
     // Popup for device diagnostics
     IF ((#hmiData.ioSlotDiagnosticsLoaded = TRUE)
       AND (#statActDeviceOfScreen >= 1)
       AND (#statActDeviceOfScreen <= "USERDIAG_DEVICES_PER_SCREEN_UPPER_LIM"))
     THEN
       #tempDeviceIndex := UINT_TO_INT(#hmiData.actIOSystemData.actIODeviceNumbers[#statActDeviceOfScreen]);
       #hmiData.actDeviceName := #ioSystemData[#statActIOSystem].devices[#tempDeviceIndex].name;
       #hmiData.actDeviceNumber := #ioSystemData[#statActIOSystem].devices[#tempDeviceIndex].number;
       #hmiData.actIPAddress := #ioSystemData[#statActIOSystem].devices[#tempDeviceIndex].ipAddress;

       FOR #tempIndex := 0 TO "USERDIAG_SLOTS_PER_SCREEN_UPPER_LIM" DO
         IF (#tempIndex <= "USERDIAG_SLOTS_PER_DEVICE_UPPER_LIM")
         THEN
           #hmiData.actIOSystemData.actDeviceSlotsUsed[#tempIndex] := (#ioSystemData[#statActIOSystem].devices[#tempDeviceIndex].slots[#tempIndex].configured);
           #hmiData.actIOSystemData.actDeviceSlotsState[#tempIndex] := #ioSystemData[#statActIOSystem].devices[#tempDeviceIndex].slots[#tempIndex].state;
         ELSE
           #hmiData.actIOSystemData.actDeviceSlotsUsed[#tempIndex] := FALSE;
           #hmiData.actIOSystemData.actDeviceSlotsState[#tempIndex] := 0;
         END_IF;
       END_FOR;
     END_IF;
     //===============================================================================================================
     // Colors the button, which switches the actual Screen of Devices in case of faulty Device is on different Screen
     //===============================================================================================================
     #tempIndex := 1;
     #tempErrorStateLower := FALSE;
     // Check if devices before the shown in actual Screen are faulty
     WHILE (#tempIndex <= (#hmiData.actIOSystemData.actIODeviceNumbers[1] - 1))
     DO
       IF ((#ioSystemData[#statActIOSystem].devices[#tempIndex].state = #STATE_FAULT)
         OR (#ioSystemData[#statActIOSystem].devices[#tempIndex].state = #STATE_LOST_CON)
         OR (#ioSystemData[#statActIOSystem].devices[#tempIndex].state = #STATE_PROBLEM))
       THEN
         #tempErrorStateLower := TRUE;
       END_IF;
       #tempIndex := #tempIndex + 1;
     END_WHILE;

     #hmiData.errorAtLowerScreen := #tempErrorStateLower;

     #tempIndex := UINT_TO_INT(#hmiData.actIOSystemData.actIODeviceNumbers["USERDIAG_DEVICES_PER_SCREEN_UPPER_LIM"] + 1);
     #tempErrorStateUpper := FALSE;
     // Check if devices after the shown in actual Screen are faulty
     IF (#tempIndex > 1)
     THEN
       WHILE ((#tempIndex <= #ioSystemData[#statActIOSystem].lastDevice))
       DO
         IF ((#ioSystemData[#statActIOSystem].devices[#tempIndex].state = #STATE_FAULT)
           OR (#ioSystemData[#statActIOSystem].devices[#tempIndex].state = #STATE_LOST_CON)
           OR (#ioSystemData[#statActIOSystem].devices[#tempIndex].state = #STATE_PROBLEM))
         THEN
           #tempErrorStateUpper := TRUE;
         END_IF;
         #tempIndex := #tempIndex + 1;
       END_WHILE;
     END_IF;

     #hmiData.errorAtUpperScreen := #tempErrorStateUpper;
     //=============================================================================
     // Check if PLC diagnostics is selected
     //=============================================================================
   ELSIF (#statActIOSystem = -1)
   THEN
     //=============================================================================
     // Acknowledge
     //=============================================================================
     IF (#hmiData.ackStates = TRUE)
     THEN
       FOR #tempIndex := 0 TO "USERDIAG_SLOTS_PER_SCREEN_UPPER_LIM" DO
         IF (#tempIndex <= "USERDIAG_SLOTS_PER_PLC_UPPER_LIM")
         THEN
           IF ((#plcData.slots[#tempIndex].state = #STATE_WAS_FAULT)
             OR (#plcData.slots[#tempIndex].state = #STATE_PROBLEM_GONE))
           THEN
             #plcData.slots[#tempIndex].state := #STATE_OK;
           END_IF;
         END_IF;
       END_FOR;
     END_IF;

     //=============================================================================
     // Copy PLC diagnostics to HMI
     //=============================================================================
     FOR #tempIndex := 0 TO "USERDIAG_SLOTS_PER_SCREEN_UPPER_LIM" DO

       IF (#tempIndex <= "USERDIAG_SLOTS_PER_PLC_UPPER_LIM")
       THEN
         #hmiData.actIOSystemData.actDeviceSlotsUsed[#tempIndex] := (#plcData.slots[#tempIndex].configured);
         #hmiData.actIOSystemData.actDeviceSlotsState[#tempIndex] := #plcData.slots[#tempIndex].state;
       ELSE
         #hmiData.actIOSystemData.actDeviceSlotsUsed[#tempIndex] := FALSE;
         #hmiData.actIOSystemData.actDeviceSlotsState[#tempIndex] := 0;
       END_IF;
     END_FOR;

   ELSE
     ; // No copy of IO System necessary
   END_IF;


   // Set Bit in HMI, if an Error occurs in IO System
   FOR #tempIoIndex := 1 TO "USERDIAG_IO_SYSTEMS_UPPER_LIM" DO
     #hmiData.ioSystemError[#tempIoIndex] := #ioSystemData[#tempIoIndex].error;
   END_FOR;
END_FUNCTION_BLOCK

// ===== PLC "_PLC"  CPU 1512SP F-1 PN =====

VAR_GLOBAL   // PLC tag table "Default tag table"
   "CARRIER_DRIVE_STATUS" AT %IW52 : Word;   // G120 D Zustandswort 1 / Stausword 1 - DRIVE / CARRIER G120 DRIVE ZSW STATUS WORD
   "CARRIER_DRIVE_WARN" AT %IW28 : Word;   // G120 D digitale Eingänge / digital Inputs - DRIVE
   "CARRIER_DRIVE_CONTROL" AT %QW300 : Word;   // G120 D Steuerwort 1 / Controlword 1 - DRIVE
   "CARRIER_DRIVE_CMD_SPEED" AT %QW302 : Word;   // G120 D Soll-Drehzahl / Setpoint-Speed of rotation - DRIVE
   "CARRIER_DRIVE_ERROR" AT %IW29 : Word;
   "HMI_IR_Remote_Control1" AT %IW200 : Word;
   "HMI_IR_Remote_Control2" AT %IW201 : Word;
   "HMI_Display_LED2" AT %QW201 : Word;
   "HMI_Display_LED1" AT %QW200 : Word;
   "HMI_Display_LED3" AT %QW202 : Word;
   "HMI_Display_DIO1_Out" AT %QW5 : Word;
   "HMI_Display_DIO1_In" AT %IW202 : Word;
   "HMI_IR_P2P" AT %IW203 : Word;
   "HMI_Device_Control" AT %IW204 : Word;
   "SpareOutput(4_7)" AT %Q4.7 : Bool;   // SPARE OUTPUT
   "Tag_3" AT %QW62 : Word;
   "temout" AT %MW0 : Word;
   "Tag_4" AT %QW250 : Word;
   "Tag_5" AT %MW200 : Word;
   "Tag_6" AT %QW161 : Word;
   "Tag_7" AT %QW162 : Word;
   "Tag_8" AT %MW2 : Word;
   "Tag_9" AT %MW52 : Word;
   "Tag_10" AT %QW280 : Word;
   "Tag_1" AT %QW2280 : Word;
   "DriveEnable" AT %M4.0 : Bool;
   "Tag_2" AT %M4.1 : Bool;
   "Tag_11" AT %QW54 : Word;
   "Tag_12" AT %QW150 : Word;
   "Tag_14" AT %QW152 : Word;
   "Drive_Status" AT %IW300 : Word;
   "TempDriveControl" AT %MW10 : Word;
   "DriveOn" AT %M4.2 : Bool;
   "Drive_Speed" AT %IW302 : Word;
   "System_Byte" AT %MB1 : Byte;
   "FirstScan" AT %M1.0 : Bool;
   "DiagStatusUpdate" AT %M1.1 : Bool;
   "AlwaysTRUE" AT %M1.2 : Bool;
   "AlwaysFALSE" AT %M1.3 : Bool;
   "Clock_Byte" AT %MB0 : Byte;
   "Clock_10Hz" AT %M0.0 : Bool;
   "Clock_5Hz" AT %M0.1 : Bool;
   "Clock_2.5Hz" AT %M0.2 : Bool;
   "Clock_2Hz" AT %M0.3 : Bool;
   "Clock_1.25Hz" AT %M0.4 : Bool;
   "Clock_1Hz" AT %M0.5 : Bool;
   "Clock_0.625Hz" AT %M0.6 : Bool;
   "Clock_0.5Hz" AT %M0.7 : Bool;
   "Running_Forward" AT %Q517.0 : Bool;
   "Running_Reverse" AT %Q517.1 : Bool;
   "Stopped" AT %Q517.2 : Bool;
   "ProductionHoldPB_Status" AT %Q517.3 : Bool;
   "CrashDetectStatus" AT %Q517.4 : Bool;
   "HeartBeat" AT %Q517.5 : Bool;
   "SDC_IN_Heartbeat" AT %I526.0 : Bool;
   "SDC_IN_Fault_Reset" AT %I526.2 : Bool;
   "Drive_Warning" AT %IW308 : Int;
   "Drive_Fault" AT %IW310 : Int;
   "AtNextStopPosition" AT %M4.3 : Bool;
   "AtPositionHighLimit" AT %MW6 : UInt;
   "AtPositionLowLimit" AT %MW8 : UInt;
   "Tag_28" AT %M90.0 : Bool;
   "SitopSelectStatus" AT %I11.3 : Bool;   // Sitop Select Status
   "DCPowerOn" AT %I11.4 : Bool;   // 24V DC Power On
   "480VPowerOn" AT %I11.5 : Bool;   // 480V DC Power On
   "Spare(11_7)" AT %I11.7 : Bool;   // Spare Input
   "Reset" AT %M2.1 : Bool;
   "SDC_IN_At_Cmd_Pos" AT %I526.3 : Bool;
   "SDC_IN_DuplicateCarrierNumber" AT %I526.4 : Bool;
   "Next_Stop_Position" AT %MW12 : UInt;
   "DuplicateCarrierFound" AT %M4.4 : Bool;
   "SDC_IN_MotionOnFault" AT %I526.5 : Bool;
   "SDC_IN_MotionOffFault" AT %I526.6 : Bool;
   "SDC_IN_CarrierSpacingFault" AT %I526.7 : Bool;
   "Tag_13" AT %I13.0 : Bool;
   "Indicon_Temp_Off" AT %M4.5 : Bool;
   "CARRIER_POSITION" AT %ID114 : DWord;
   "DisconnectOn" AT %I11.0 : Bool;   // Disconnect On
   "SpareInput(11_2)" AT %I11.2 : Bool;   // Spare Input
   "ProductionHoldPB_LH" AT %I12.0 : Bool;   // Production Hold Button LH
   "ResetPB_LH" AT %I12.1 : Bool;   // Reset Push Button LH
   "ProductionHoldPB_RH" AT %I12.2 : Bool;   // Production Hold Button RH
   "ResetPB_RH" AT %I12.3 : Bool;   // Reset Push Button RH
   "Spare(12_4)" AT %I12.4 : Bool;   // Spare Input
   "Spare(12_5)" AT %I12.5 : Bool;   // Spare Input
   "Spare(12_6)" AT %I12.6 : Bool;   // Spare Input
   "Spare(12_7)" AT %I12.7 : Bool;   // Spare Input
   "FaultLight_RH" AT %Q4.3 : Bool;   // FAULT LIGHT RH
   "RunLight_LH" AT %Q4.2 : Bool;   // RUN LIGHT LH
   "FaultLight_LH" AT %Q4.1 : Bool;   // FAULT LIGHT LH
   "IRD400_HMI_24VDC_ENABLE" AT %Q4.0 : Bool;   // IRD 400 PANEL HMI 24V DC POWER
   "RunLight_RH" AT %Q4.4 : Bool;   // RUN LIGHT RH
   "SpareOutput(4_6)" AT %Q4.6 : Bool;   // SPARE OUTPUT
   "SpareOutput(4_5)" AT %Q4.5 : Bool;   // SPARE OUTPUT
   "SpareSafetyOutput(6_7)" AT %Q6.7 : Bool;   // SPARE SAFETY OUTPUT
   "SpareSafetyOutput(6_6)" AT %Q6.6 : Bool;   // SPARE SAFETY OUTPUT
   "SpareSafetyOutput(6_5)" AT %Q6.5 : Bool;   // SPARE SAFETY OUTPUT
   "SpareSafetyOutput(6_4)" AT %Q6.4 : Bool;   // SPARE SAFETY OUTPUT
   "Crash_Detect_OK(6)" AT %Q6.3 : Bool;   // SPARE SAFETY OUTPUT
   "SpareSafetyOutput(6_2)" AT %Q6.2 : Bool;   // SPARE SAFETY OUTPUT
   "SpareSafetyOutput(6_1)" AT %Q6.1 : Bool;   // SPARE SAFETY OUTPUT
   "Crash_Detect_OK" AT %Q6.0 : Bool;   // Carrier Crash Detect
   "Slot3_SafetyOutput" AT %QW6 : Word;
   "Slot2_SafetyInput" AT %IW0 : Word;
   "Slot4_Input" AT %IW11 : Word;
   "Slot5_Output" AT %QW4 : Word;
   "CARRIER01_POSITION_SDC_OUT" AT %QD512 : DWord;
   "SectionComment" AT %M4.6 : Bool;
   "EncoderERR" AT %I110.0 : Bool;
   "EncoderWRN" AT %I110.1 : Bool;
   "EncoderNP" AT %I110.2 : Bool;
   "EncoderEV" AT %I110.3 : Bool;
   "EncoderYPosition" AT %ID116 : DWord;
   "EncoderXPosition" AT %ID112 : DWord;
   "Crash_Detect_Prox" AT %I11.6 : Bool;   // Spare Input
   "EncoderErrorCode" AT %IW114 : Word;
   "Accumulator_PE" AT %I11.1 : Bool;   // Spare Input
END_VAR

VAR_GLOBAL   // PLC tag table "To_SDC_TagTable"
   "ToSDC_Status" AT %QW510 : Word;   // CARRIER STATUS WORD
   "ToSDC_Status.0" AT %Q510.0 : Bool;   // HEARTBEAT
   "ToSDC_Status.1" AT %Q510.1 : Bool;   // MANUAL
   "ToSDC_Status.2" AT %Q510.2 : Bool;   // IN_AUTO
   "ToSDC_Status.3" AT %Q510.3 : Bool;   // POSITIONING_COMPLETE
   "ToSDC_Status.4" AT %Q510.4 : Bool;   // PRODUCTION HOLD
   "ToSDC_Status.5" AT %Q510.5 : Bool;   // CARRIER MOVING FORWARD
   "ToSDC_Status.6" AT %Q510.6 : Bool;   // CARRIER MOVING REVERSE
   "ToSDC_Status.7" AT %Q510.7 : Bool;   // CARRIER FAULT
   "ToSDC_Status.8" AT %Q511.0 : Bool;   // CRASH DETECT TRIPPED
   "ToSDC_Status.9" AT %Q511.1 : Bool;   // ENCODER COMM FAULT
   "ToSDC_Status.10" AT %Q511.2 : Bool;   // DRIVE COMM FAULT
   "ToSDC_Status.11" AT %Q511.3 : Bool;   // HMI COMM FAULT
   "ToSDC_Status.12" AT %Q511.4 : Bool;
   "ToSDC_Status.13" AT %Q511.5 : Bool;
   "ToSDC_Status.14" AT %Q511.6 : Bool;
   "ToSDC_Status.15" AT %Q511.7 : Bool;
   "ToSDC_FaultCode" AT %QW512 : Word;   // SDC FAULT CODE
   "ToSDC_CarrierPosition" AT %QD514 : DWord;   // CARRIER POSITION
   "ToSDC_CarrierNumber" AT %QW518 : Word;   // CARRIER NUMBER
   "ToSDC_G120DControlWord" AT %QW520 : Word;   // G120D_STW1_CONTROL
   "ToSDC_G120DControlWord.0" AT %Q520.0 : Bool;   // Bit_00_ON
   "ToSDC_G120DControlWord.1" AT %Q520.1 : Bool;   // Bit_01_AUS2_INH
   "ToSDC_G120DControlWord.2" AT %Q520.2 : Bool;   // Bit_02_AUS3_STOP
   "ToSDC_G120DControlWord.3" AT %Q520.3 : Bool;   // Bit_03_EN
   "ToSDC_G120DControlWord.4" AT %Q520.4 : Bool;   // Bit_04_EN_RAMP
   "ToSDC_G120DControlWord.5" AT %Q520.5 : Bool;   // Bit_05_START_RAMP
   "ToSDC_G120DControlWord.6" AT %Q520.6 : Bool;   // Bit_06_SETPOINT
   "ToSDC_G120DControlWord.7" AT %Q520.7 : Bool;   // Bit_07_RESET
   "ToSDC_G120DControlWord.8" AT %Q521.0 : Bool;   // Bit_08_JOG_R
   "ToSDC_G120DControlWord.9" AT %Q521.1 : Bool;   // Bit_09_JOG_L
   "ToSDC_G120DControlWord.10" AT %Q521.2 : Bool;   // Bit_10_CONTR_PLC
   "ToSDC_G120DControlWord.11" AT %Q521.3 : Bool;   // Bit_11_REVERSE
   "ToSDC_G120DControlWord.12" AT %Q521.4 : Bool;   // Bit_12_BRAKE_RELEASE
   "ToSDC_G120DControlWord.13" AT %Q521.5 : Bool;   // Bit_13_DDS
   "ToSDC_G120DControlWord.14" AT %Q521.6 : Bool;   // Bit_14_DO0
   "ToSDC_G120DControlWord.15" AT %Q521.7 : Bool;   // Bit_15_DO1
   "ToSDC_G120DStatusWORD" AT %QW522 : Word;   // G120D_ZSW1_STATUS
   "ToSDC_G120DStatusWORD.0" AT %Q522.0 : Bool;   // Bit_00_READY_RUN
   "ToSDC_G120DStatusWORD.1" AT %Q522.1 : Bool;   // Bit_01_READY_ON
   "ToSDC_G120DStatusWORD.2" AT %Q522.2 : Bool;   // Bit_02_ENABLE
   "ToSDC_G120DStatusWORD.3" AT %Q522.3 : Bool;   // Bit_03_FAULT
   "ToSDC_G120DStatusWORD.4" AT %Q522.4 : Bool;   // Bit_04_OFF2
   "ToSDC_G120DStatusWORD.5" AT %Q522.5 : Bool;   // Bit_05_OFF3
   "ToSDC_G120DStatusWORD.6" AT %Q522.6 : Bool;   // Bit_06_LOCK_OUT
   "ToSDC_G120DStatusWORD.7" AT %Q522.7 : Bool;   // Bit_07_WARN
   "ToSDC_G120DStatusWORD.8" AT %Q523.0 : Bool;   // Bit_08_NO_DEVIATION
   "ToSDC_G120DStatusWORD.9" AT %Q523.1 : Bool;   // Bit_09_CONTR_PLC
   "ToSDC_G120DStatusWORD.10" AT %Q523.2 : Bool;   // Bit_10_F_MAX
   "ToSDC_G120DStatusWORD.11" AT %Q523.3 : Bool;   // Bit_11_LIMIT_REACHED
   "ToSDC_G120DStatusWORD.12" AT %Q523.4 : Bool;   // Bit_12_BRAKE_OPEN
   "ToSDC_G120DStatusWORD.13" AT %Q523.5 : Bool;   // Bit_13_NO_OVERTEMP
   "ToSDC_G120DStatusWORD.14" AT %Q523.6 : Bool;   // Bit_14_CW_CCW
   "ToSDC_G120DStatusWORD.15" AT %Q523.7 : Bool;   // Bit_15_OVERL
   "ToSDC_Slot2Input" AT %QB524 : Byte;   // SLOT 2 INPUT WORD
   "ToSDC_CrashDetectSW" AT %Q524.0 : Bool;   // CRASH DETECT SW
   "ToSDC_SpareSafetyInput(21)" AT %Q524.1 : Bool;   // SPARE SAFETY INPUT
   "ToSDC_SpareSafetyInput(22)" AT %Q524.2 : Bool;   // SPARE SAFETY INPUT
   "ToSDC_SpareSafetyInput(23)" AT %Q524.3 : Bool;   // SPARE SAFETY INPUT
   "ToSDC_SpareSafetyInput(24)" AT %Q524.4 : Bool;   // SPARE SAFETY INPUT
   "ToSDC_SpareSafetyInput(25)" AT %Q524.5 : Bool;   // SPARE SAFETY INPUT
   "ToSDC_SpareSafetyInput(26)" AT %Q524.6 : Bool;   // SPARE SAFETY INPUT
   "ToSDC_SpareSafetyInput(27)" AT %Q524.7 : Bool;   // SPARE SAFETY INPUT
   "ToSDC_Slot3SafetyOutput" AT %QB525 : Byte;   // SLOT 3 SAFETY OUTPUT WORD
   "ToSDC_CrashDetectOK" AT %Q525.0 : Bool;   // CARRIER CRASH DETECT
   "ToSDC_SpareSafetyOutput(31)" AT %Q525.1 : Bool;   // SPARE SAFETY OUTPUT
   "ToSDC_SpareSafetyOutput(32)" AT %Q525.2 : Bool;   // SPARE SAFETY OUTPUT
   "ToSDC_SpareSafetyOutput(33)" AT %Q525.3 : Bool;   // SPARE SAFETY OUTPUT
   "ToSDC_SpareSafetyOutput(34)" AT %Q525.4 : Bool;   // SPARE SAFETY OUTPUT
   "ToSDC_SpareSafetyOutput(35)" AT %Q525.5 : Bool;   // SPARE SAFETY OUTPUT
   "ToSDC_SpareSafetyOutput(36)" AT %Q525.6 : Bool;   // SPARE SAFETY OUTPUT
   "ToSDC_SpareSafetyOutput(37)" AT %Q525.7 : Bool;   // SPARE SAFETY OUTPUT
   "ToSDC_Slot4Input" AT %QW526 : Word;   // SLOT 4 INPUT WORD
   "ToSDC_480VPowerOnMDCB1" AT %Q526.0 : Bool;   // 480 VAC POWER ON MDCB 1
   "ToSDC_SpareInput(41)" AT %Q526.1 : Bool;   // SPARE INPUT
   "ToSDC_SpareInput(42)" AT %Q526.2 : Bool;   // SPARE INPUT
   "ToSDC_SitopSelectStatus" AT %Q526.3 : Bool;   // SITOP SELECT STATUS
   "ToSDC_DCsupplyOnPSCB2" AT %Q526.4 : Bool;   // DC SUPPLY ON PSCB 2
   "ToSDC_SpareInput(45)" AT %Q526.5 : Bool;   // SPARE INPUT
   "ToSDC_SpareInput(46)" AT %Q526.6 : Bool;   // SPARE INPUT
   "ToSDC_SpareInput(47)" AT %Q526.7 : Bool;   // SPARE INPUT
   "ToSDC_PB1ProdHoldLH" AT %Q527.0 : Bool;   // PB 1 PRODUCTION HOLD LH
   "ToSDC_PB2ResetLH" AT %Q527.1 : Bool;   // PB 2 RESET LH
   "ToSDC_PB3ProdHoldRH" AT %Q527.2 : Bool;   // PB 3 PRODUCTION HOLD RH
   "ToSDC_PB4ResetRH" AT %Q527.3 : Bool;   // PB 4 RESET RH
   "ToSDC_SpareInput(414)" AT %Q527.4 : Bool;   // SPARE INPUT
   "ToSDC_SpareInput(415)" AT %Q527.5 : Bool;   // SPARE INPUT
   "ToSDC_SpareInput(416)" AT %Q527.6 : Bool;   // SPARE INPUT
   "ToSDC_SpareInput(417)" AT %Q527.7 : Bool;   // SPARE INPUT
   "ToSDC_Slot5Output" AT %QB528 : Byte;   // SLOT 5 OUTPUT WORD
   "ToSDC_IRD400HMI24VDCENABLE" AT %Q528.0 : Bool;   // IRD 400 PANEL HMI 24V DC POWER
   "ToSDC_FaultLightLH" AT %Q528.1 : Bool;   // FAULT LIGHT LH
   "ToSDC_RunLightLH" AT %Q528.2 : Bool;   // RUN LIGHT LH
   "ToSDC_FaultLightRH" AT %Q528.3 : Bool;   // FAULT LIGHT RH
   "ToSDC_RunLightRH" AT %Q528.4 : Bool;   // RUN LIGHT RH
   "ToSDC_SpareOutput(55)" AT %Q528.5 : Bool;   // SPARE OUTPUT
   "ToSDC_SpareOutput(56)" AT %Q528.6 : Bool;   // SPARE OUTPUT
   "ToSDC_SpareOutput(57)" AT %Q528.7 : Bool;   // SPARE OUTPUT
   "ToSDC_ActualSpeed" AT %QW530 : Word;   // ACTUAL SPEED
   "ToSDC_CarrierDriveAlarm" AT %QW532 : Word;   // CARRIER DRIVE ALARM
   "ToSDC_CarrierDriveWarning" AT %QW534 : Word;   // CARRIER DRIVE WARNING
END_VAR

VAR_GLOBAL   // PLC tag table "From_SDC_TagTable"
   "FromSDC_CarrierInZone" AT %IW510 : Word;
   "FromSDC_CarrierNumberEcho" AT %IW512 : Word;
   "FromSDC_CarrierPositionEcho" AT %ID514 : DWord;
   "FromSDC_NextCarriernumber" AT %IW518 : Word;
   "FromSDC_Nextstopposition" AT %ID520 : DWord;
   "FromSDC_DriveCommandSpeed" AT %IW524 : Word;
   "FromSDC_DuplicateCarrierNumber" AT %IW526 : Word;
   "FromSDC_FirstDuplicateCarrierPosition" AT %ID528 : DWord;
   "FromSDC_SecondDuplicateCarrierPosition" AT %ID532 : DWord;
   "FromSDC_CommandWord" AT %IW536 : Word;
   "FromSDC_Heartbeat" AT %I536.0 : Bool;
   "FromSDC_DriveForwardCommand" AT %I536.1 : Bool;
   "FromSDC_FaultReset" AT %I536.2 : Bool;
   "FromSDC_AtCommandPosition" AT %I536.3 : Bool;
   "FromSDC_DuplicateCarrierFault" AT %I536.4 : Bool;
   "FromSDC_MotionOnFault" AT %I536.5 : Bool;
   "FromSDC_MotionOffFault" AT %I536.6 : Bool;
   "FromSDC_CarrierSpacingFault" AT %I536.7 : Bool;
END_VAR

TYPE "UDT_Carrier"
VERSION : 0.1
   STRUCT
      Position : DWord;
      CarrierNumber : Word;
      CarrierInZone : Word;
      ActualSpeed : Word;   // Drive Speed in Hz
      Stopped : Bool;
      MovingFwd : Bool;
      MovingRev : Bool;
      Ready : Bool;
      ReadyOn : Bool;
      Enabled : Bool;
      Fault : Bool;
      CollisionAlarm : Bool;
      Encoder : "UDT_PnF_Pxv_Encoder";
      DriveControl : "UDT_G120D_STW1_CONTROL";
      DriveStatus : "UDT_G120D_ZSW1_STATUS";
      Error : "UDT_G120D_ERRORS";
      CommandSpeed : Word;
      ProductionHold : Bool;
      Reset : Bool;
      NextCarrierNum : Word;
      NextCarrierPos : Word;
      HMI : "UDT_CarrierHMI";
      IR_Remote : "UDT_IRD400";
      SDC_IN : "UDT_SDC_IN";
      SDC_Out : "UDT_SDC_OUT";
      JOG : "UDT_Jog";
      Semi_Auto : "UDT_SEMI_AUTO";
      Mode : "UDT_Mode";
      LH_PB_Box : "UDT_PB_Box";
      RH_PB_Box : "UDT_PB_Box";
   END_STRUCT;
END_TYPE

TYPE "UDT_EMS"
VERSION : 0.1
   STRUCT
      CARRIER : Array[1..99] of "UDT_Carrier";
   END_STRUCT;
END_TYPE

TYPE "UDT_CarrierHMI_In"
   STRUCT
      JogFWD : Bool;
      JogRev : Bool;
      FaultStatus : Array[0..20] of Bool;
      ResetFault : Bool;
   END_STRUCT;
END_TYPE

TYPE "UDT_ZONE"
   STRUCT
      ZONE : Int;
      START_POSITION : Int;
      STOP_POSITION : Int;
      DESCRIPTION : String;
   END_STRUCT;
END_TYPE

TYPE "UDT_CarrierHMI_Out"
   STRUCT
      Faults : Bool;
   END_STRUCT;
END_TYPE

TYPE "UDT_CarrierHMI"
   STRUCT
      HMI_In : "UDT_CarrierHMI_In";
      HMI_Out : "UDT_CarrierHMI_Out";
   END_STRUCT;
END_TYPE

TYPE "UDT_SDC_OUT"
   STRUCT
      CarrierNumber : Word;
      CarrierPosition : Word;
      ActualSpeed : Word;
      CarrierDriveFaults : Word;
      CarrierDriveAlarms : Word;
      CarrierFaults : Word;
      Spare_Word : Word;
      RunningFWD : Bool;
      RunningREV : Bool;
      Stopped : Bool;
      ProductionHoldPB_Status : Bool;
      CrashDetectStatus : Bool;
      HeartBeat : Bool;
      AutoMode : Bool;
      ManualMode : Bool;
   END_STRUCT;
END_TYPE

TYPE "UDT_SDC_IN"
   STRUCT
      Zone : Int;
      CarrierNumEcho : Word;
      CarrierPositionEcho : DWord;
      NextCarrierNum : Word;
      NextStopPos : DWord;
      DriveFwdCMD : Bool;
      DriveCmdSpeed : Word;
      Spare_Word_1 : Word;
      Spare_Word_2 : Word;
      HeartBeat : Bool;
      FaultReset : Bool;
      HighSpeedEnable : Bool;
      AtCmdPos : Bool;
      DuplicateCarrierNumber : Int;
      FirstDuplicateCarrierPosition : Word;
      SecondDuplicateCarrierPosition : Word;
      Faults : "UDT_SDC_IN_FAULTS";
   END_STRUCT;
END_TYPE

TYPE "UDT_PnF_Pxv_EncoderPositionModule"
   STRUCT
      XPos : DWord;
      YPos : DWord;
   END_STRUCT;
END_TYPE

TYPE "GF_Zeit_Messung"
VERSION : 0.1
   STRUCT
      akt : Int;   // Zeitwert in Mykrosekunden
      min : Int;   // Zeitwert in Mykrosekunden
      max : Int;   // Zeitwert in Mykrosekunden
      Speicher : LReal;   // Zwischenspeicher
   END_STRUCT;
END_TYPE

TYPE "UDT_MAIN"
   STRUCT
      AlwaysOn : Bool;
      AutoMode : Bool;
      ManualMode : Bool;
   END_STRUCT;
END_TYPE

TYPE "UDT_IRD400"
   STRUCT
      Segment1 : Byte;
      Segment2 : Byte;
      Segment3 : Byte;
      DisplayLED : Byte;
      DisplayControl : Byte;
      F1_Key : Bool;
      F2_Key : Bool;
      PL_Key : Bool;
      "(*)_Key" : Bool;
      Enter_Key : Bool;
      ESC : Bool;
      "1_Key" : Bool;
      "2_Key" : Bool;
      "3_Key" : Bool;
      "4_Key" : Bool;
      "5_Key" : Bool;
      "6_Key" : Bool;
      "7_Key" : Bool;
      "8_Key" : Bool;
      "9_Key" : Bool;
      "0_Key" : Bool;
   END_STRUCT;
END_TYPE

TYPE "UDT_Jog"
VERSION : 0.1
   STRUCT
      JogFWDFast : Bool;
      JogFWDMed : Bool;
      JogFWDSlow : Bool;
      JogREVFast : Bool;
      JogREVMed : Bool;
      JogREVSlow : Bool;
      JogSpeedSlow : Word;
      JogSpeedMed : Word;
      JogSpeedFast : Word;
      JogCommand : Bool;
   END_STRUCT;
END_TYPE

TYPE "UDT_Mode"
   STRUCT
      AutoMode : Bool;
      ManualMode : Bool;
      ManualMode_Enable : Bool;
      SemiAutoMode : Bool;
      IR_First_Number : String;
      IR_Second_Number : String;
      IR_Third_Number : String;
      IR_First_Two_Digits : String;
      IR_Number_Entered : String[3];
      IR_First_Number_Null : Bool;
      IR_Second_Number_Null : Bool;
      IR_Third_Number_Null : Bool;
      IR_Any_Number_Pressed : Bool;
      IR_First_Number_ONS : Bool;
      IR_Second_Number_ONS : Bool;
      IR_Third_Number_ONS : Bool;
      IR_Number_Entered_INT : Int;
   END_STRUCT;
END_TYPE

TYPE "UDT_SDC_IN_FAULTS"
   STRUCT
      DuplicateCarrierFault : Bool;
      MotionOnFault : Bool;
      MotionOffFault : Bool;
      CarrierSpacingFault : Bool;
   END_STRUCT;
END_TYPE

TYPE "UDT_SEMI_AUTO"
   STRUCT
      MoveToNxtStpEnable : Bool;   // Move To Next in Manual Mode
      MoveToNxtStpAntiRep : Bool;   // Move to Next Stop Manual Mode Anti Repeat
      MoveToNxtStpAntiRepRst : Bool;   // Move to Next Stop Manual Mode Anti Repeat Reset
   END_STRUCT;
END_TYPE

TYPE "UDT_PB_Box_Out"
   STRUCT
      SafetySolenoid : Bool;
      SitopReset : Bool;
      FaultLT : Bool;
      RunLT : Bool;
      ProdHoldLT : Bool;
   END_STRUCT;
END_TYPE

TYPE "UDT_PB_Box"
   STRUCT
      In : "UDT_PB_Box_In";
      Out : "UDT_PB_Box_Out";
   END_STRUCT;
END_TYPE

TYPE "UDT_PB_Box_In"
   STRUCT
      Crash_Detect_SW : Bool;
      "480VAC_PowerOn" : Bool;
      SitopSelectStatus : Bool;
      DC_PowerOn : Bool;
      ProdHold : Bool;
      ResetPB : Bool;
   END_STRUCT;
END_TYPE

TYPE "UDT_PnF_Pxv_Encoder"
   STRUCT
      PositionMod : "UDT_PnF_Pxv_EncoderPositionModule";
      Position : DWord;
      StatusMod : "UDT_PnF_Pxv_EncoderStatusModule";
   END_STRUCT;
END_TYPE

TYPE "UDT_PnF_Pxv_EncoderStatusModule"
   STRUCT
      Status : Word;
      Error : Bool;
      NoPosition : Bool;
      Warning : Bool;
      Event : Bool;
      ErrorCode : Word;
   END_STRUCT;
END_TYPE

TYPE "UDT_G120D_STW1_CONTROL"
VERSION : 0.1
   STRUCT
      Bit_08_JOG_R : Bool;   // 1=tippen rechtsseitig EIN/ 0= AUS / 1=jogging on right-hand side ON/ 0= OFF
      Bit_09_JOG_L : Bool;   // 1=tippen linksseitig EIN/ 0= AUS / 1=jogging on left-hand side ON/ 0= OFF
      Bit_10_CONTR_PLC : Bool;   // 1=Bedienung über PLC erforderlich/ 0=keine Bedienung über PLC erforderlich / 1=control by PLC required/ 0=no control by PLC required
      Bit_11_REVERSE : Bool;   // 1=Umkehrung des Sollwerts/ 0=keine Umkehrung / 1=inversion of setpoint/ 0=no inversion of setpoint
      Bit_12_BRAKE_Release : Bool;   // 1= Löse Bremse / 1= Release Break / 1= Manual Brake Release
      Bit_13_DDS : Bool;   // 1=DDS1 FU Datenset / 0=DDS0 FU Datenset / 1=DDS1 FU Dataset / 0=DDS0 FU Dataset
      Bit_14_DO0 : Bool;   // 1=Digitaler Ausgang aktiv/ 0=Digitaler Ausgang nicht aktiv / 1=Digital Output activ/ 0=Digital Output not activ
      Bit_15_DO1 : Bool;   // 1=Digitaler Ausgang aktiv/ 0=Digitaler Ausgang nicht aktiv / 1=Digital Output activ/ 0=Digital Output not activ
      Bit_00_ON : Bool;   // 1=EIN/ 0=AUS / 1=ON/ 0=OFF2
      Bit_01_AUS2_INH : Bool;   // 1=Betriebsvoraussetzung/ 0=AUS2 - Pulsverzögerer, Spannung auf einmal aus / 1=operation condition/ 0=AUS2 - pulse inhibitor, voltage off at once
      Bit_02_AUS3_STOP : Bool;   // 1=Betriebsvoraussetzung / 0=AUS3 - schneller Halt / 1=operation condition / 0=AUS3 - fast stop
      Bit_03_EN : Bool;   // 1=Freigabe Betrieb/ 0=deaktiviere Betrieb / 1=enable operation/ 0=disable operation
      Bit_04_EN_RAMP : Bool;   // 1=1=Betriebsvoraussetzung / 0=deaktiviere Funktionsrampengenerator / 1=operation condition / 0=disable ramp function generator
      Bit_05_START_RAMP : Bool;   // 1=Aktiviere Rampenfunktion / 0=deaktivere RFG / 1=enable ramp function generator / 0=stoppen RFG
      Bit_06_SETPOINT : Bool;   // 1=Freigabe Sollwert/ 0=deaktiviere Sollwert / 1=enable setpoint/ 0=disable setpoint
      Bit_07_RESET : Bool;   // 1=Störung quittieren / 0= irrelevant / 1=Reset fault / 0= irrelevant
   END_STRUCT;
END_TYPE

TYPE "UDT_G120D_ZSW1_STATUS"
VERSION : 0.1
   STRUCT
      Bit_08_NO_DEVIATION : Bool;   // 1=keine Abweichung des Sollwerts / 0=Abweichung / 1=no deviation current-setpoint / 0=deviation / Setpoint / actual value deviation within the tolerance range.
      Bit_09_CONTR_PLC : Bool;   // 1=Kontrolle über PLC erforderlich/ 0=keine Kontrolle erforderlich / 1=control by PLC required/ 0=no control by PLC required / The automation system is requested to ac-cept the inverter control.
      Bit_10_F_MAX : Bool;   // 1=fmax erreicht/ 0= unter fmax / 1=fmax reached/ 0= below fmax / Speed is greater than or equal to the corre-sponding maximum speed.
      Bit_11_LIMIT_REACHED : Bool;   // 1=keine Warnung/ 0=Warnung: Motor an Spannungsgrenze / 1=no warning/ 0=warning:Motor at limit of current / Comparison value for current or torque has been reached or exceeded.
      Bit_12_BRAKE_OPEN : Bool;   // 1= / 0=Haltebremse / motor Brake is open
      Bit_13_NO_OVERTEMP : Bool;   // 1= / 0=Motorüberlast / Drive Overtemperature
      Bit_14_CW_CCW : Bool;   // 1=Rechtslauf/ 0=Linkslauf / On for drive runnin clockwise/off counterclockwise
      Bit_15_OVERL : Bool;   // 1= /0= Konvertierer Überlast / 1= /0= Konverter overload / 0 = Alarm, in-verter thermal overload/on CDS display
      Bit_00_READY_RUN : Bool;   // 1=bereit zum betreiben/ 0= nicht bereit / 1=ready to run/ 0= not ready to run / Power supply switched on; electronics initial-ized; pulses locked.
      Bit_01_READY_ON : Bool;   // 1=bereit zum einschalten/ 0= nicht bereit / 1=ready to switch on/ 0= not ready to switch on / Motor is switched on (ON/OFF1 = 1), no fault is active. With the command "Enable opera-tion" (STW1.3), the inverter switches on the motor.
      Bit_02_ENABLE : Bool;   // 1=Freigabe Bedienung / 0=deaktiviere Bedienung / 1=operation enabled / 0=operation disabled / Motor follows setpoint. See control word 1, bit 3.
      Bit_03_FAULT : Bool;   // 1=Störung / 0=keine Störung / 1=fault / 0=no fault / The inverter has a fault. Acknowledge fault using STW1.7
      Bit_04_OFF2 : Bool;   // 1=kein AUS2 / 0=AUS2 Befehl ist vorhanden / 1=no AUS2 / 0=AUS2 command is present / OFF2 Coast down to standstill is not active.
      Bit_05_OFF3 : Bool;   // 1=kein AUS3 / 0=AUS3 Befehl ist vorhanden / 1=no AUS3 / 0=AUS3 command is present / OFF3 Quick stop is not active.
      Bit_06_LOCK_OUT : Bool;   // 1=sperre Ausschaltung / 0=keine Sperrung / 1=closing lock-out / 0=no closing lock-out / It is only possible to switch on the motor after an OFF1 followed by ON.
      Bit_07_WARN : Bool;   // 1=Warnung / 0= keine Warnung / 1=Warning / 0= no warning
   END_STRUCT;
END_TYPE

TYPE "UDT_G120D_ERRORS"
VERSION : 0.1
   STRUCT
      F_X33_F1 : Bool;   // Fehler Überstrom / Fault Overcurrent / Overcurrent
      F_X34_F2 : Bool;   // Fehler Überspannung / Fault Overvoltage / Overvoltage
      F_X35_F3 : Bool;   // Fehler Unterspannung / Fault Undervoltage / Undervoltage
      F_X36_F4 : Bool;   // Fehler Inverter Übertemperatur / Fault Inverter over temperature / Motor Data recognition fault
      F_X37_F41 : Bool;   // Fehler Motordatenerkennung / Motor data identification failure / Motor Data recognition fault
      F_X38_F52 : Bool;   // Fehler Leistungsteil / Power stack Fault / Error Power Section
      F_X39_F62 : Bool;   // Fehler MMC Daten sind fehlerhaft / Fault MMC contents invalid / Error MCC data is faulty
      F_X40_F70 : Bool;   // Fehler PLC Sollposition / PLC setpoint fault
      F_X41_F71 : Bool;   // Fehler USS Sollposition, Überwachung / USS setpoint fault, monitoring
      F_X42_F72 : Bool;   // Fehler USS Sollposition, USS Master / USS setpoint fault, USS master
      F_X43_F90 : Bool;   // Fehler Gebersignal / Faulty encoder signal
      F_X44_F395 : Bool;   // Fehler CU/PM wechsel / Fault CU/PM swap
      bit_14 : Bool;   // Reserve / spare
      bit_15 : Bool;   // Reserve / spare
      bit_16 : Bool;   // Reserve / spare
      bit_17 : Bool;   // Reserve / spare
   END_STRUCT;
END_TYPE

DATA_BLOCK "Main_Safety_RTG1_DB"   // DB1, F_DB
{ S7_Optimized_Access := 'TRUE' }
NAME : FUSI
VERSION : 0.1
"Main_Safety_RTG1"
BEGIN
END_DATA_BLOCK

// folder: 05_DB'S

DATA_BLOCK "FB_G120D_DB"   // DB2
{ S7_Optimized_Access := 'FALSE' }
VERSION : 0.1
"FB105_G120D_CarrierDrive"
BEGIN
END_DATA_BLOCK

DATA_BLOCK "Default_SupervisionDB"   // DB3
{ S7_Optimized_Access := 'TRUE' }
VERSION : 0.1
"FB1000_Default_SupervisionFB"
BEGIN
END_DATA_BLOCK

DATA_BLOCK "LSitop_PseDiag_DB"   // DB12
{ S7_Optimized_Access := 'FALSE' }
AUTHOR : DFCS
FAMILY : SITOP
VERSION : 2.3
"LSitop_PseDiag"
BEGIN
END_DATA_BLOCK

DATA_BLOCK "InstAGV"   // DB14
{ S7_Optimized_Access := 'TRUE' }
AUTHOR : Siemens
VERSION : 1.0
"FB104_CarrierBreakerStatus"
BEGIN
END_DATA_BLOCK

DATA_BLOCK "Global"   // DB15
{ S7_Optimized_Access := 'TRUE' }
AUTHOR : Siemens
VERSION : 1.0
   VAR
      MyLadder : Hw_Device := 32;
      MyMode : UInt := 0;
      ReturnValue : Int;
      MyState : Array[0..127] of Bool;
      System : Struct   // Functiongroup system
         Diagnosis : Struct   // System diagnosis
            Fuse : Struct
               Channel1 : Bool;   // Channel 1 active
               Channel2 : Bool;   // Channel 2 active
               Channel3 : Bool;   // Channel 3 active
               Channel4 : Bool;   // Channel 4 active
               CollectiveError : Bool;   // Collective error sensitivity module
            END_STRUCT;
            Profinet : Struct
               CollectiveError : Bool;   // Collective error Profinet IO
               Status : Array[0..1023] of Bool;   // Device status disturbed
            END_STRUCT;
            Profibus : Struct
               CollectiveError : Bool;   // Collective error Profibus DP
            END_STRUCT;
         END_STRUCT;
      END_STRUCT;
   END_VAR
BEGIN
END_DATA_BLOCK

DATA_BLOCK "CARRIER"   // DB100
{ S7_Optimized_Access := 'TRUE' }
VERSION : 0.1
BEGIN
END_DATA_BLOCK

DATA_BLOCK "DB101_CARRIER_CONTROL"   // DB101
{ S7_Optimized_Access := 'TRUE' }
VERSION : 0.1
   VAR
      CARRIER_CONTROL_IN : "UDT_G120D_STW1_CONTROL";
   END_VAR
BEGIN
END_DATA_BLOCK

DATA_BLOCK "SYSTEM"   // DB104
{ S7_Optimized_Access := 'TRUE' }
VERSION : 0.1
   VAR
      MAIN : "UDT_MAIN";
   END_VAR
BEGIN
END_DATA_BLOCK

DATA_BLOCK "SDC_IN"   // DB110
{ S7_Optimized_Access := 'TRUE' }
VERSION : 0.1
   VAR
      Input : "UDT_SDC_OUT";
   END_VAR
BEGIN
END_DATA_BLOCK

DATA_BLOCK "SDC_OUT"   // DB111
{ S7_Optimized_Access := 'TRUE' }
VERSION : 0.1
   VAR
      Output : "UDT_SDC_IN";
   END_VAR
BEGIN
END_DATA_BLOCK

DATA_BLOCK "DB300_FAULTS"   // DB300
{ S7_Optimized_Access := 'TRUE' }
VERSION : 0.1
   VAR
      Faults : Word;
   END_VAR
BEGIN
END_DATA_BLOCK

DATA_BLOCK "DB1110_Red_Green_LED"   // DB1110
{ S7_Optimized_Access := 'TRUE' }
VERSION : 0.1
"FB1110_Red_Green_LED"
BEGIN
   instWRREC.LEN := 1;
END_DATA_BLOCK

// folder: 06_IDBs

DATA_BLOCK "FB_Carrier_DB"   // DB6
{ S7_Optimized_Access := 'TRUE' }
VERSION : 0.1
"FB100_Carrier"
BEGIN
END_DATA_BLOCK

DATA_BLOCK "Decode_Carrier_Number_DB"   // DB16
{ S7_Optimized_Access := 'TRUE' }
VERSION : 0.1
"FB103_Decode_Carrier_Number"
BEGIN
END_DATA_BLOCK

DATA_BLOCK "Decode_Speed_DB"   // DB17
{ S7_Optimized_Access := 'TRUE' }
VERSION : 0.1
"FB102_Decode_Speed"
BEGIN
END_DATA_BLOCK

// folder: 08_SYSTEM

DATA_BLOCK "VS"   // DB250
TITLE = System- Variablen
{ S7_Optimized_Access := 'TRUE' }
VERSION : 0.1
// Allgem. Variablen wie z.B. ZTakte, VKE_0 usw.,
// die im ges. Programm (auch innerhalb von MModul-Bausteinen) ausgewertet werden. Ein Beschreiben dieser Variablen ist nicht zulässig.
// Variablen dürfen auch nicht an Ausgangs/ oder Ein/Ausgangsparameter parametriert werden.
   VAR
      "Takt_0,1s" : Bool;   // Taktmerker 10 Hz
      "Takt_0,2s" : Bool;   // Taktmerker 5 Hz
      "Takt_0,4s" : Bool;   // Taktmerker 2,5 Hz
      "Takt_0,5s" : Bool;   // Taktmerker 2 Hz
      "Takt_0,8s" : Bool;   // Taktmerker 1,25 Hz
      "Takt 1s" : Bool;   // Taktmerker 1Hz
      "Takt_1,6s" : Bool;   // Taktmerker 0,625 Hz
      Takt_2s : Bool;   // Taktmerker 0,5 Hz
      "ZTakt_0,1s" : Bool;   // Zähltakt 0,1s
      ZTakt_1s : Bool;   // Zähltakt 1s
      "Trig_0,1s" : Bool;   // Triggermerker Zähltakt 0,1s
      BliS : Bool;   // Blinktakt schnell
      BliL : Bool;   // Blinktakt langsam
      Anl_Verlae : Bool;   // Anlauf verlängert (während Resetzeit)
      Neustart : Bool;   // Neustart
      "Reset-Init" : Bool;   // Reset-Init manuelle Ansteuerung
      "Resst-Init-Imp" : Bool;   // Reset-Init-Impuls für 1Zyklus
      "Reset-Ein" : Bool;   // Reset- Impuls für 1 Zyklus bei Steuerung Ein
      Reset : Bool;   // Reset-Impuls bei Steuerung 1 über Zeit
      Steu_ein : Bool;
      VKE0 : Bool;   // VKE0 für prov. Unterbrechungen
      VKE1 : Bool;   // VKE1 für prov. Brücken
      Null : Bool;   // Null-Merker für Parametrierungen
      Eins : Bool;   // Eins-Merker für Parametrierungen
      Mit : Bool;   // Mit-Merker für Auswahlen
      Ohne : Bool;   // Ohne-Merker für Auswahlen
      "??????" : Bool;   // Platzhalter
      Dunkel : Bool;   // Dunkelschaltung
      Mel_int : Bool;   // Melderkontrolle intern
      Kon_int : Bool;   // Kontrollen intern
      Sifa_int : Bool;   // Sicherungsfall intern
      AQu_EnStoe : Bool;   // automatische Störungsquittung
      AQu_UeZeit : Bool;   // automatische Überwachungszeitnachtriggerung
      Allg_Stoe : Bool;   // Allgemeine Störungen
      PN_Fehler : Bool;   // Profinetstörung
      S_K0 : Bool;   // Steuerung Ein an Sicherheitsprog.
      F_ZykZeit : Bool;   // Anzeige Zykluszeitfehler
      F_DiagAlarm : Bool;   // Anzeige diagnosefähige Baugruppe defekt
      F_BG_Wechsel : Bool;   // Anzeige Baugruppe raus / rein / Kontaktfehler
      F_BG_Ausfall : Bool;   // Anzeige Baugruppenträger Ausfall
      F_ProgFehler : Bool;   // Anzeige Programmfehler
      F_Periph_Zugr : Bool;   // Anzeige Fehler beim Peripherie-Zugriff
   END_VAR
BEGIN
END_DATA_BLOCK

DATA_BLOCK "01_GrFunkt_DB"   // DB500
{ S7_Optimized_Access := 'TRUE' }
VERSION : 0.1
"01_GrFunkt"
BEGIN
END_DATA_BLOCK

DATA_BLOCK "GF_An_Vor_St"   // DB501
{ S7_Optimized_Access := 'TRUE' }
VERSION : 0.1
   VAR RETAIN
      Res : Array[1..8] of Byte;   // Reserve
      max_Anzahl : Int := 40;   // maximale Anzahl der An/Vorwahlen
   END_VAR
BEGIN
END_DATA_BLOCK

DATA_BLOCK "GF_BetrArt_St"   // DB502
{ S7_Optimized_Access := 'TRUE' }
VERSION : 0.1
   VAR RETAIN
      Res : Array[1..8] of Byte;   // Reserve
      max_Anzahl : Int := 20;   // maximale Anzahl der Betriebsarten
   END_VAR
BEGIN
END_DATA_BLOCK

DATA_BLOCK "GF_Grund_DB"   // DB503
{ S7_Optimized_Access := 'TRUE' }
AUTHOR : Audi
FAMILY : Grund
NAME : Grund_DB
VERSION : 2.0
   VAR RETAIN
      Akt_Datum_Uhrzeit : DTL := DTL#2014-03-18-14:56:01.55;   // Aktuelle Datum / Uhrzeit von AG
      Akt_Datum_Uhrzeit_ASCII : Struct   // Aktuelle Datum / Uhrzeit von AG
         Datum : Struct   // Datum
            Jahr : Array[1..4] of Char;   // Jahr
            Monat : Array[1..2] of Char;   // Monat
            Tag : Array[1..2] of Char;   // Tag
            YYYYMMDD : String[8];   // Datum Format YYYYMMDD
         END_STRUCT;
         Zeit : Struct   // Zeit
            Stunde : Array[1..2] of Char;   // Stunde
            Minute : Array[1..2] of Char;   // Minute
            Sekunde : Array[1..2] of Char;   // Sekunde
            MilliSek : Array[1..3] of Char;   // Milisekunde
            HHMMSS : String[6];   // Zeit Format hhmmss
         END_STRUCT;
         Wochentag : Char := '3';
      END_STRUCT;
      Stellbits : Struct
         Stell_ASCII : Bool := false;   // Stellbit von LAN-Paket
         Stell_OPs : Bool := false;   // Stellbit an OP's
         OP_Stell : Bool := false;   // Stellbit von OP
      END_STRUCT;
   END_VAR
   VAR
      Stell_Datum_Uhrzeit : DTL := DTL#1970-01-01-00:00:00;   // AG-Stell Datum / Uhrzeit
   END_VAR
   VAR RETAIN
      Stell_Datum_Uhrzeit_ASCI : Struct   // AG_Stell Datum / Uhrzeit
         Jahr : Array[1..4] of Char;
         Monat : Array[1..2] of Char;
         Tag : Array[1..2] of Char;
         Stunde : Array[1..2] of Char;
         Minute : Array[1..2] of Char;
         Sekunde : Array[1..2] of Char;
         MilliSek : Array[1..3] of Char;
         Wochentag : Char := ' ';
      END_STRUCT;
      Ret_Val : Int;
      Anlagenname : String[8];
      Reserve : Array[1..4] of Byte;
      Zyklusstatistik : Struct
         System : Struct
            akt_Zykluszeit : Int := 0;   // aktuelle Zykluszeit OB1
            min_Zykluszeit : Int := 0;   // minimale Zykluszeit OB1
            max_Zykluszeit : Int := 0;   // minimale Zykluszeit OB1
         END_STRUCT;
         gem_min_Zykluszeit : Int := 0;   // gemessene minimale Zykluszeit
         gem_max_Zykluszeit : Int := 0;   // gemessene maximale Zykluszeit
         Zeit_SichProg : Int := 0;   // Zeit Ablauf Sicherheitsprogramm
         Res_Gem_ZyklZeit : Bool := false;   // Reset gemessene Zykluszeit
         Reserve : String[2] := '';
      END_STRUCT;
   END_VAR
   VAR
      Res_Zeit : Array[1..10] of Bool;
      Zeit : Array[1..10] of "GF_Zeit_Messung";
      ZLT : Struct
         Anwahl_mit_ZLT : Bool;
         "akt_S-Punkt" : Struct
            Z_Pkt : String[4];   // Zeitpunkt (erste Zeit)
            S_Info : String[2];   // Schaltinformation
            S_Info_hex : Byte;   // Schaltinformation in hex
         END_STRUCT;
         "nächst_S-Punkt" : Struct
            Z_Pkt : String[4];   // Zeitpunkt (erste Zeit)
            S_Info : String[2];   // Schaltinformation
         END_STRUCT;
         Geschw_ZLT : Int;
         Geschw_Man : Int;
         Akt_Geschw : Int;
         Zeit : Array[1..6] of Char;
         Datum : Array[1..6] of Char;
         Zeit_hhmm : Array[1..4] of Char;
      END_STRUCT;
      Zeit_Ma_PC : String[24];   // Zeitformat Master-PC YYYY-MM-TT__hh:mm:ss:mmm
   END_VAR
BEGIN
   Stell_Datum_Uhrzeit_ASCI.Jahr[1] := ' ';
   Stell_Datum_Uhrzeit_ASCI.Jahr[2] := ' ';
   Stell_Datum_Uhrzeit_ASCI.Jahr[3] := ' ';
   Stell_Datum_Uhrzeit_ASCI.Jahr[4] := ' ';
   Stell_Datum_Uhrzeit_ASCI.Monat[1] := ' ';
   Stell_Datum_Uhrzeit_ASCI.Monat[2] := ' ';
   Stell_Datum_Uhrzeit_ASCI.Tag[1] := ' ';
   Stell_Datum_Uhrzeit_ASCI.Tag[2] := ' ';
   Stell_Datum_Uhrzeit_ASCI.Stunde[1] := ' ';
   Stell_Datum_Uhrzeit_ASCI.Stunde[2] := ' ';
   Stell_Datum_Uhrzeit_ASCI.Minute[1] := ' ';
   Stell_Datum_Uhrzeit_ASCI.Minute[2] := ' ';
   Stell_Datum_Uhrzeit_ASCI.Sekunde[1] := ' ';
   Stell_Datum_Uhrzeit_ASCI.Sekunde[2] := ' ';
   Stell_Datum_Uhrzeit_ASCI.MilliSek[1] := ' ';
   Stell_Datum_Uhrzeit_ASCI.MilliSek[2] := ' ';
   Stell_Datum_Uhrzeit_ASCI.MilliSek[3] := ' ';
   Reserve[1] := 16#00;
   Reserve[2] := 16#00;
   Reserve[3] := 16#00;
   Reserve[4] := 16#00;
   Akt_Datum_Uhrzeit_ASCII.Datum.Jahr[1] := '2';
   Akt_Datum_Uhrzeit_ASCII.Datum.Jahr[2] := '0';
   Akt_Datum_Uhrzeit_ASCII.Datum.Jahr[3] := '1';
   Akt_Datum_Uhrzeit_ASCII.Datum.Jahr[4] := '4';
   Akt_Datum_Uhrzeit_ASCII.Datum.Monat[1] := ' ';
   Akt_Datum_Uhrzeit_ASCII.Datum.Monat[2] := '3';
   Akt_Datum_Uhrzeit_ASCII.Datum.Tag[1] := '1';
   Akt_Datum_Uhrzeit_ASCII.Datum.Tag[2] := '8';
   Akt_Datum_Uhrzeit_ASCII.Zeit.Stunde[1] := '1';
   Akt_Datum_Uhrzeit_ASCII.Zeit.Stunde[2] := '4';
   Akt_Datum_Uhrzeit_ASCII.Zeit.Minute[1] := '5';
   Akt_Datum_Uhrzeit_ASCII.Zeit.Minute[2] := '6';
   Akt_Datum_Uhrzeit_ASCII.Zeit.Sekunde[1] := ' ';
   Akt_Datum_Uhrzeit_ASCII.Zeit.Sekunde[2] := '1';
   Akt_Datum_Uhrzeit_ASCII.Zeit.MilliSek[1] := '5';
   Akt_Datum_Uhrzeit_ASCII.Zeit.MilliSek[2] := '5';
   Akt_Datum_Uhrzeit_ASCII.Zeit.MilliSek[3] := '0';
END_DATA_BLOCK

DATA_BLOCK "GF_HBed_Obj_St"   // DB504
{ S7_Optimized_Access := 'TRUE' }
VERSION : 0.1
   VAR RETAIN
      Res : Array[1..8] of Byte;   // Reserve
      max_Anzahl : Int := 299;   // maximale Anzahl der An/Vorwahlen
   END_VAR
BEGIN
END_DATA_BLOCK

DATA_BLOCK "GF_LastSp_St"   // DB506
{ S7_Optimized_Access := 'TRUE' }
VERSION : 0.1
   VAR RETAIN
      Zentr_EinAus : Struct   // Zentrale Ein/Ausschaltung der Lastspannung
         AnwZLT : Bool;   // Anwahl ZLT-Betrieb
         EinZ : Bool;   // Ein von ZLT
         Ausz : Bool;   // Aus von ZLT
         EinS : Bool;   // Ein von Schalktschrank
         AusS : Bool;   // Aus von Schaltschrank
      END_STRUCT;
      Res : Array[1..6] of Byte;   // Reserve
      max_Anzahl : Int := 20;   // maximale Anzahl der Lastspannungen
   END_VAR
BEGIN
END_DATA_BLOCK

DATA_BLOCK "GF_Visu_allg"   // DB507
{ S7_Optimized_Access := 'TRUE' }
VERSION : 0.1
   VAR
      AAE : Struct   // Anzeige Analogwerte-Energie
         Frg_Anwahl : Bool;   // Freigabe Werte-Auswahl
         Pult : String[4];   // Pultname das ausgewählt hat
         A_Anwahl : Int;   // Auswahl
      END_STRUCT;
   END_VAR
   VAR RETAIN
      Test_WS : Int;
   END_VAR
   VAR
      Test_St : Struct
         Test_2 : Int;
      END_STRUCT;
   END_VAR
BEGIN
END_DATA_BLOCK

DATA_BLOCK "PN_DiagDB"   // DB508
{ S7_Optimized_Access := 'FALSE' }
AUTHOR : Audi
FAMILY : Profibus
NAME : PB_DiagD
VERSION : 1.0
   VAR
      vonVisu : Struct
         HMI_ID : Word;   // Nr. des OP, welches den DB benutzt (0 = unbenutzt)
         IOSys_ID : Int;   // von Visu angef. IO-System-ID 1 od. 2 = PB; 100 od. 101 =PN
         TLN_Nr : Int;   // Teilnehmer-Nr
         Res : DWord;
      END_STRUCT;
      PN100 : Struct
         S_Bereich : Array[1..32] of Struct   // Störbereich
            Stoe : Bool;   // Störmeldung
            TN_Beginn : Int;   // 1.Teilnehmer für Zusammenfassung Störbereich
            TN_Ende : Int;   // letzter Teilnehmer Zusammenfassung Störbereich
         END_STRUCT;
         res : Array[1..8] of Byte;
         konfig_TN : Array[0..1023] of Bool;   // Mode_1: Bitleiste für alle im Master parametrierten Teilnehmer
         fehlerhafte_TN : Array[0..1023] of Bool;   // Bitleiste für alle fehlerhaften Teilnehmer
         gestörte_TN : Array[0..1023] of Bool;   // Mode_2: Bitleiste für alle gestörten Teilnehmer
         deaktiviert_TN : Array[0..1023] of Bool;   // Mode_3: Bitleiste für alle deaktivierten Teilnehmer
         vorhanden_TN : Array[0..1023] of Bool;   // Mode_4: Bitleiste für alle vorhandenen Teilnehmer
         problem_TN : Array[0..1023] of Bool;   // Mode_5: Bitleiste für alle Teilnehmer mit einem Problem
      END_STRUCT;
      Reserve : String[4];
   END_VAR
BEGIN
   PN100.S_Bereich[1].TN_Beginn := 1;
   PN100.S_Bereich[1].TN_Ende := 5;
   PN100.S_Bereich[2].TN_Beginn := 6;
   PN100.S_Bereich[2].TN_Ende := 10;
   PN100.S_Bereich[3].TN_Beginn := 11;
   PN100.S_Bereich[3].TN_Ende := 120;
END_DATA_BLOCK

DATA_BLOCK "PN_Zykl_DB"   // DB509
{ S7_Optimized_Access := 'FALSE' }
AUTHOR : Audi
FAMILY : Profibus
NAME : PB_Zykl
VERSION : 1.0
"PN_Zykl"
BEGIN
END_DATA_BLOCK

// folder: System blocks/Program resources

DATA_BLOCK "SDC_Heartbeat_On_Timer"   // DB4
{ S7_Optimized_Access := 'TRUE' }
AUTHOR : Simatic
FAMILY : IEC
NAME : IEC_TMR
VERSION : 1.0
"IEC_TIMER"
BEGIN
END_DATA_BLOCK

DATA_BLOCK "SDC_Heartbeat_Off_Timer"   // DB11
{ S7_Optimized_Access := 'TRUE' }
AUTHOR : Simatic
FAMILY : IEC
NAME : IEC_TMR
VERSION : 1.0
"IEC_TIMER"
BEGIN
END_DATA_BLOCK

// folder: (top level)

FUNCTION_BLOCK "Main_Safety_RTG1"   // FB0, F_FBD
{ S7_Optimized_Access := 'TRUE' }
VERSION : 0.1
BEGIN
END_FUNCTION_BLOCK

ORGANIZATION_BLOCK "Main"   // OB1, LAD, ProgramCycle
TITLE = "Main Program Sweep (Cycle)"
{ S7_Optimized_Access := 'FALSE' }
VERSION : 0.1
   VAR_TEMP
      EV_CLASS : Byte;   // Bits 0-3 = 1:Coming event, Bits 4-7 = 1:Event class 1
      SCAN_1 : Byte;   // 1:Initial call of the OB, 3: Call 2-n of the OB
      PRIORITY : Byte;   // Priority of OB Execution
      OB_NUMBR : Byte;   // OB number
      RESERVED_1 : Byte;   // Reserved for system
      RESERVED_2 : Byte;   // Reserved for system
      PREV_CYCLE : Int;   // Previous program cycle time (milliseconds)
      MIN_CYCLE : Int;   // Minimum program cycle time (milliseconds)
      MAX_CYCLE : Int;   // Maximum program cycle time (milliseconds)
      DATE_TIME : Date_And_Time;   // Date and time OB started
      tempreceive : Word;
   END_VAR
BEGIN

REGION Network 1
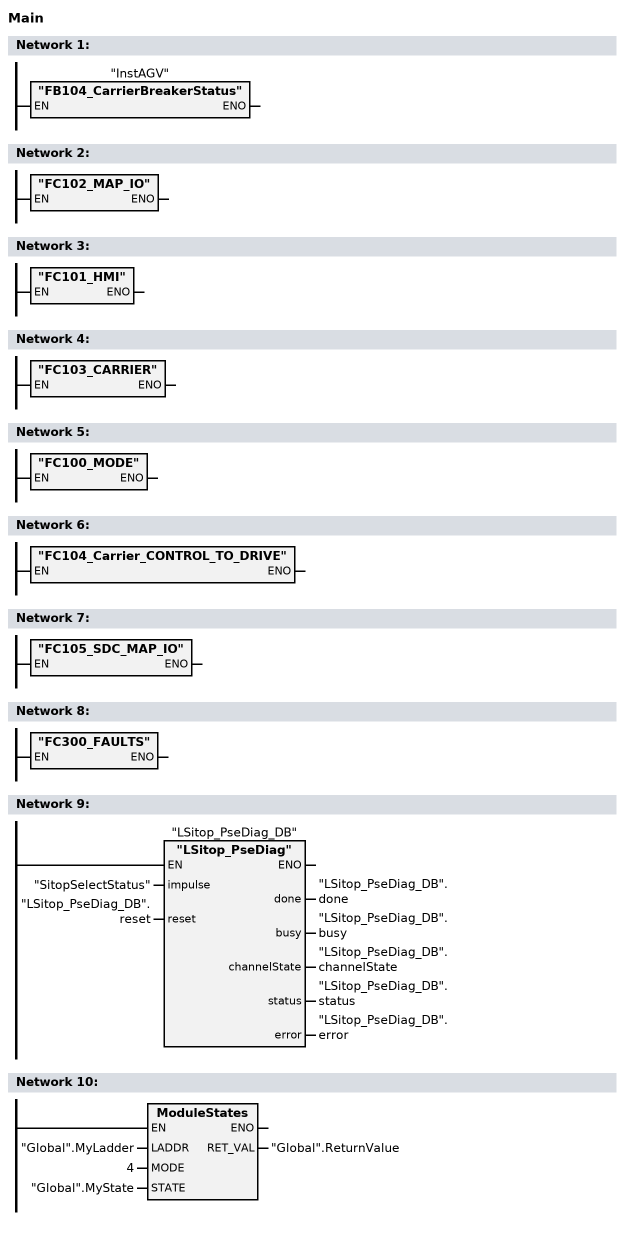
   RUNG wire#powerrail
      "InstAGV"()
   END_RUNG
   // the same network as SCL:
   "InstAGV"();   // "FB104_CarrierBreakerStatus"
END_REGION

REGION Network 2
   RUNG wire#powerrail
      "FC102_MAP_IO"()
   END_RUNG
   // the same network as SCL:
   "FC102_MAP_IO"();
END_REGION

REGION Network 3
   RUNG wire#powerrail
      "FC101_HMI"()
   END_RUNG
   // the same network as SCL:
   "FC101_HMI"();
END_REGION

REGION Network 4
   RUNG wire#powerrail
      "FC103_CARRIER"()
   END_RUNG
   // the same network as SCL:
   "FC103_CARRIER"();
END_REGION

REGION Network 5
   RUNG wire#powerrail
      "FC100_MODE"()
   END_RUNG
   // the same network as SCL:
   "FC100_MODE"();
END_REGION

REGION Network 6
   RUNG wire#powerrail
      "FC104_Carrier_CONTROL_TO_DRIVE"()
   END_RUNG
   // the same network as SCL:
   "FC104_Carrier_CONTROL_TO_DRIVE"();
END_REGION

REGION Network 7
   RUNG wire#powerrail
      "FC105_SDC_MAP_IO"()
   END_RUNG
   // the same network as SCL:
   "FC105_SDC_MAP_IO"();
END_REGION

REGION Network 8
   RUNG wire#powerrail
      "FC300_FAULTS"()
   END_RUNG
   // the same network as SCL:
   "FC300_FAULTS"();
END_REGION

REGION Network 9
   RUNG wire#powerrail
      "LSitop_PseDiag_DB"(impulse := "SitopSelectStatus", reset := "LSitop_PseDiag_DB".reset, done => "LSitop_PseDiag_DB".done, busy => "LSitop_PseDiag_DB".busy, channelState => "LSitop_PseDiag_DB".channelState, status => "LSitop_PseDiag_DB".status, error => "LSitop_PseDiag_DB".error)
   END_RUNG
   // the same network as SCL:
   "LSitop_PseDiag_DB"(impulse := "SitopSelectStatus",   // "LSitop_PseDiag"
                       reset := "LSitop_PseDiag_DB".reset,
                       done => "LSitop_PseDiag_DB".done,
                       busy => "LSitop_PseDiag_DB".busy,
                       channelState => "LSitop_PseDiag_DB".channelState,
                       status => "LSitop_PseDiag_DB".status,
                       error => "LSitop_PseDiag_DB".error);
END_REGION

REGION Network 10
   // no SCL statement known for ModuleStates: written as a call
   "Global".ReturnValue := ModuleStates(LADDR := "Global".MyLadder, MODE := 4, STATE := "Global".MyState);
END_REGION
END_ORGANIZATION_BLOCK

ORGANIZATION_BLOCK "ProDiagOB"   // OB250, ProDiag_OB, ProgramCycle
TITLE = "Main Program Sweep (Cycle)"
{ S7_Optimized_Access := 'TRUE' }
VERSION : 0.1
   VAR_INPUT
      Initial_Call : Bool;   // Initial call of this OB
      Remanence : Bool;   // =True, if remanent data are available
   END_VAR
BEGIN

REGION Network 1
   CALL "FB1000_Default_SupervisionFB", "Default_SupervisionDB";
END_REGION
END_ORGANIZATION_BLOCK

// folder: 03_FB'S

